// TIA Portal project "CHEMICAL DOSING PUMP" (V16)

(* hardware
DEVICE "S7-1200 station_1"  S7-1200 Station
   slot 0: "Rack_0"  S7-1200 Rack  Rack  V1.0
   slot 1: "PLC_1"  CPU 1214C DC/DC/DC  6ES7 214-1AG40-0XB0  V4.4
DEVICE "HMI_1"  TP900 Comfort
   slot 0: "HMI_1"  TP900 Comfort  6AV2 124-0JC01-0AX0  16.0.0.0
   slot 1: "HMI_RT_1"  TP900 Comfort  6AV2 124-0JC01-0AX0  16.0.0.0
   slot 5: "HMI_1.IE_CP_1"  PROFINET Interface  16.0.0.0
      slot 1: "PROFINET Interface_1"  PROFINET Interface
         slot 1: "Port_1"  Port
         slot 2: "Port_2"  Port
   slot 7: "HMI_1.MPI/DP_CP_1"  MPI/DP Interface  16.0.0.0
*)

// ===== PLC "PLC_1"  CPU 1214C DC/DC/DC =====

VAR_GLOBAL   // PLC tag table "Default tag table"
   "STOP SYSTEM" AT %M0.0 : Bool;
   "START SYSTEM" AT %M0.1 : Bool;
   "SYSTEM RUNNING" AT %M0.2 : Bool;
   "System_Byte" AT %MB2000 : Byte;
   "FirstScan" AT %M2000.0 : Bool;
   "DiagStatusUpdate" AT %M2000.1 : Bool;
   "AlwaysTRUE" AT %M2000.2 : Bool;
   "AlwaysFALSE" AT %M2000.3 : Bool;
   "System_Byte(1)" AT %MB1 : Byte;
   "Clock_Byte" AT %MB2001 : Byte;
   "Clock_10Hz" AT %M2001.0 : Bool;
   "Clock_5Hz" AT %M2001.1 : Bool;
   "Clock_2.5Hz" AT %M2001.2 : Bool;
   "Clock_2Hz" AT %M2001.3 : Bool;
   "Clock_1.25Hz" AT %M2001.4 : Bool;
   "Clock_1Hz" AT %M2001.5 : Bool;
   "Clock_0.625Hz" AT %M2001.6 : Bool;
   "Clock_0.5Hz" AT %M2001.7 : Bool;
   "TRIGGER 1" AT %M0.3 : Bool;
   "TRIGGER 2" AT %M0.4 : Bool;
   "DOSING PUMP 1" AT %Q0.0 : Bool;
   "HIGH LEVEL SET POINT" AT %MW4 : Int;
   "WATER TANK 2" AT %MW2 : Int;
   "TRIGGER 3" AT %M0.5 : Bool;
   "DOSING PUMP 2" AT %Q0.1 : Bool;
   "WATER TANK 2_2" AT %MW6 : Int;
   "TRIGGER 4" AT %M0.6 : Bool;
   "TRIGGER 5" AT %M0.7 : Bool;
   "TRIGGER 6" AT %M1.0 : Bool;
   "LOW LEVEL SETPOINT" AT %MW8 : Int;
END_VAR

// folder: System blocks/Program resources

DATA_BLOCK "C0"   // DB1
{ S7_Optimized_Access := 'TRUE' }
AUTHOR : Simatic
FAMILY : IEC
NAME : CNTR
VERSION : 1.0
// stored: InstanceOfName IEC_COUNTER
"IEC_COUNTER"
BEGIN
END_DATA_BLOCK

DATA_BLOCK "C1"   // DB2
{ S7_Optimized_Access := 'TRUE' }
AUTHOR : Simatic
FAMILY : IEC
NAME : CNTR
VERSION : 1.0
// stored: InstanceOfName IEC_COUNTER
"IEC_COUNTER"
BEGIN
END_DATA_BLOCK

// folder: (top level)

ORGANIZATION_BLOCK "Main"   // OB1, LAD, ProgramCycle
TITLE = "Main Program Sweep (Cycle)"
{ S7_Optimized_Access := 'TRUE' }
VERSION : 0.1
   VAR_INPUT
      Initial_Call : Bool;   // Initial call of this OB
      Remanence : Bool;   // =True, if remanent data are available
   END_VAR
   VAR_TEMP   // added for the SCL form of the ladder/FBD networks
      _w1 : Bool;
      _w2 : Bool;
      _w3 : Bool;
      _w4 : Bool;
   END_VAR
BEGIN

REGION Network 1: PROGRAM FOT STARTING AND STOPING A SYSTEM
   // * CREATING PROGRAM FOR STARTING AND STOPING CHEICAL DOSING SYSTEM
   // * ENABILY THE CLOCK MEMORY
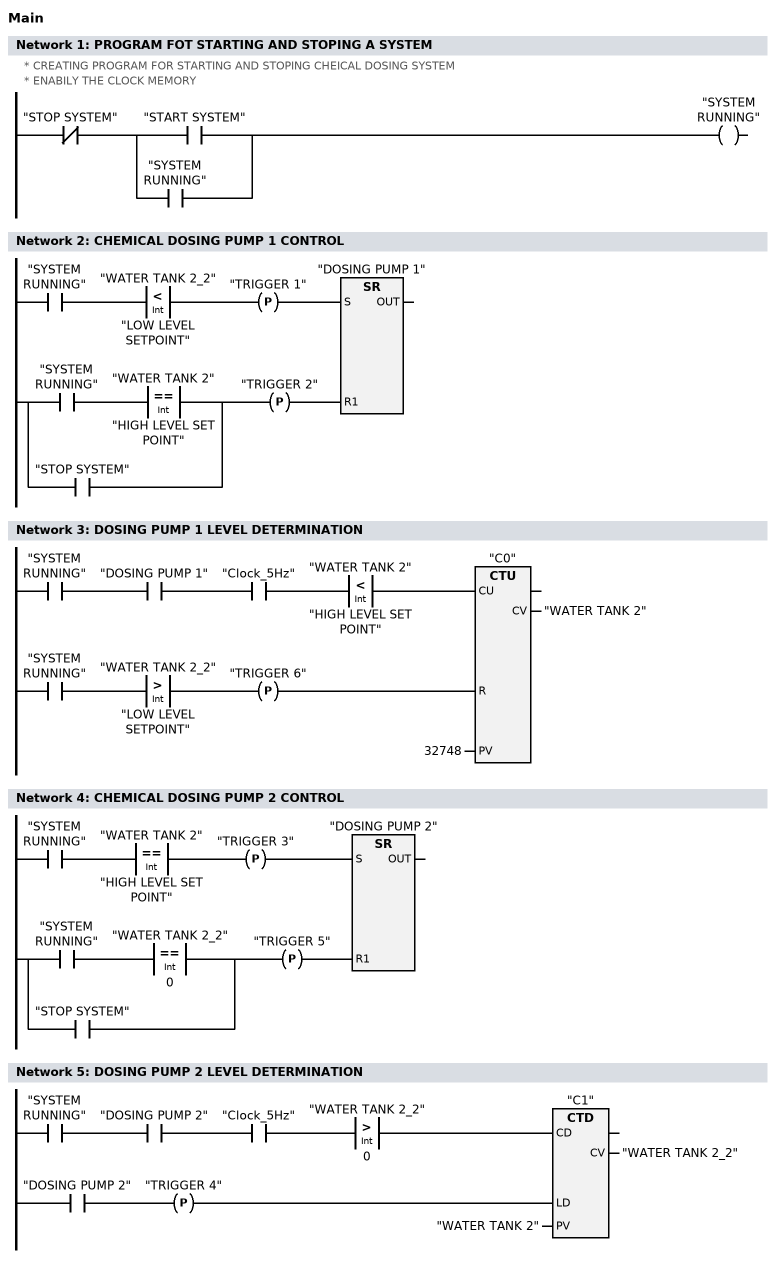
   RUNG wire#powerrail
      I_Contact( "STOP SYSTEM" )
      wire#w1
      Contact( "START SYSTEM" )
      wire#w2
      Coil( "SYSTEM RUNNING" )
   END_RUNG
   RUNG wire#w1
      Contact( "SYSTEM RUNNING" )
   END_RUNG wire#w2
   // the same network as SCL:
   "SYSTEM RUNNING" := NOT "STOP SYSTEM" AND ("START SYSTEM" OR "SYSTEM RUNNING");
END_REGION

REGION Network 2: CHEMICAL DOSING PUMP 1 CONTROL
   RUNG wire#powerrail
      Contact( "SYSTEM RUNNING" )
      { S7_Templates := "SrcType := Int" } LT_Contact(in1 := "WATER TANK 2_2", in2 := "LOW LEVEL SETPOINT")
      P_Trig( "TRIGGER 1" )
      S_SR(operand := "DOSING PUMP 1", r1 := wire#w2)
   END_RUNG
   RUNG wire#powerrail
      Contact( "SYSTEM RUNNING" )
      { S7_Templates := "SrcType := Int" } EQ_Contact(in1 := "WATER TANK 2", in2 := "HIGH LEVEL SET POINT")
      wire#w1
      P_Trig( "TRIGGER 2" )
   END_RUNG wire#w2
   RUNG wire#powerrail
      Contact( "STOP SYSTEM" )
   END_RUNG wire#w1
   // the same network as SCL:
   #_w1 := "SYSTEM RUNNING" AND ("WATER TANK 2_2" < "LOW LEVEL SETPOINT");
   #_w2 := #_w1 AND NOT "TRIGGER 1";   // rising edge
   "TRIGGER 1" := #_w1;
   #_w3 := ("SYSTEM RUNNING" AND ("WATER TANK 2" = "HIGH LEVEL SET POINT")) OR "STOP SYSTEM";
   #_w4 := #_w3 AND NOT "TRIGGER 2";   // rising edge
   "TRIGGER 2" := #_w3;
   IF #_w2 THEN
       "DOSING PUMP 1" := TRUE;   // SR flip-flop
   END_IF;
   IF #_w4 THEN "DOSING PUMP 1" := FALSE; END_IF;
END_REGION

REGION Network 3: DOSING PUMP 1 LEVEL DETERMINATION
   #_w1 := "SYSTEM RUNNING" AND ("WATER TANK 2_2" > "LOW LEVEL SETPOINT");
   #_w2 := #_w1 AND NOT "TRIGGER 6";   // rising edge
   "TRIGGER 6" := #_w1;
   "C0".CTU(CU := "SYSTEM RUNNING" AND "DOSING PUMP 1" AND "Clock_5Hz" AND ("WATER TANK 2" < "HIGH LEVEL SET POINT"),
            R := #_w2,
            PV := 32748,
            CV => "WATER TANK 2");
END_REGION

REGION Network 4: CHEMICAL DOSING PUMP 2 CONTROL
   RUNG wire#powerrail
      Contact( "SYSTEM RUNNING" )
      { S7_Templates := "SrcType := Int" } EQ_Contact(in1 := "WATER TANK 2", in2 := "HIGH LEVEL SET POINT")
      P_Trig( "TRIGGER 3" )
      S_SR(operand := "DOSING PUMP 2", r1 := wire#w2)
   END_RUNG
   RUNG wire#powerrail
      Contact( "SYSTEM RUNNING" )
      { S7_Templates := "SrcType := Int" } EQ_Contact(in1 := "WATER TANK 2_2", in2 := 0)
      wire#w1
      P_Trig( "TRIGGER 5" )
   END_RUNG wire#w2
   RUNG wire#powerrail
      Contact( "STOP SYSTEM" )
   END_RUNG wire#w1
   // the same network as SCL:
   #_w1 := "SYSTEM RUNNING" AND ("WATER TANK 2" = "HIGH LEVEL SET POINT");
   #_w2 := #_w1 AND NOT "TRIGGER 3";   // rising edge
   "TRIGGER 3" := #_w1;
   #_w3 := ("SYSTEM RUNNING" AND ("WATER TANK 2_2" = 0)) OR "STOP SYSTEM";
   #_w4 := #_w3 AND NOT "TRIGGER 5";   // rising edge
   "TRIGGER 5" := #_w3;
   IF #_w2 THEN
       "DOSING PUMP 2" := TRUE;   // SR flip-flop
   END_IF;
   IF #_w4 THEN "DOSING PUMP 2" := FALSE; END_IF;
END_REGION

REGION Network 5: DOSING PUMP 2 LEVEL DETERMINATION
   #_w1 := "DOSING PUMP 2" AND NOT "TRIGGER 4";   // rising edge
   "TRIGGER 4" := "DOSING PUMP 2";
   "C1".CTD(CD := "SYSTEM RUNNING" AND "DOSING PUMP 2" AND "Clock_5Hz" AND ("WATER TANK 2_2" > 0),
            LD := #_w1,
            PV := "WATER TANK 2",
            CV => "WATER TANK 2_2");
END_REGION
END_ORGANIZATION_BLOCK

(* ===== HMI "HMI_RT_1" =====
system functions are stored by id; their names below are inferred from use
connection "HMI_Connection_1": ETHERNET, S7_1200_OMS

HMI tags "Default tag table"
   "Tag_ScreenNumber" : UInt, internal
   "WATER TANK 2" : Int = PLC "WATER TANK 2" AT %MW2, 1 s
   "WATER TANK 2_2" : Int = PLC "WATER TANK 2_2" AT %MW6, 1 s
   "START SYSTEM" : Bool = PLC "STOP SYSTEM" AT %M0.0, 1 s
   "STOP SYSTEM" : Bool = PLC "START SYSTEM" AT %M0.1, 1 s
   "DOSING PUMP 1" : Bool = PLC "DOSING PUMP 1" AT %Q0.0, 1 s
   "DOSING PUMP 2" : Bool = PLC "DOSING PUMP 2" AT %Q0.1, 1 s
   "LOW LEVEL SETPOINT" : Int = PLC "LOW LEVEL SETPOINT" AT %MW8, 1 s
   "HIGH LEVEL SET POINT" : Int = PLC "HIGH LEVEL SET POINT" AT %MW4, 1 s
   "SYSTEM RUNNING" : Bool = PLC "SYSTEM RUNNING" AT %M0.2, 1 s

screen "Root screen" 800x420, template "Template_1"
   on GenerateScreen: SetTag("Tag_ScreenNumber", 1)
   SymbolLibrary "Symbol library_1" at 626,75 size 164x120
      Appearance <- "DOSING PUMP 1"
   SymbolLibrary "Symbol library_2" at 36,242 size 187x102
      Appearance <- "DOSING PUMP 2"
   SymbolLibrary "Symbol library_3" at 503,134 size 127x35
      Appearance <- "DOSING PUMP 1"
   SymbolLibrary "Symbol library_4" at 446,134 size 60x68
      Appearance <- "DOSING PUMP 1"
   SymbolLibrary "Symbol library_5" at 446,200 size 31x82
      Appearance <- "DOSING PUMP 1"
   SymbolLibrary "Symbol library_9" at 627,11 size 41x67
      Appearance <- "DOSING PUMP 1"
   SymbolLibrary "Symbol library_10" at 222,278 size 52x46
      Appearance <- "DOSING PUMP 2"
   SymbolLibrary "Symbol library_11" at 248,193 size 26x94
      Appearance <- "DOSING PUMP 2"
   SymbolLibrary "Symbol library_12" at 159,209 size 39x37
      Appearance <- "DOSING PUMP 2"
   SymbolLibrary "Symbol library_13" at 27,208 size 138x21
      Appearance <- "DOSING PUMP 2"
   Bar "Bar_2" at 52,76 size 280x126; MinimumValue 0; MaximumValue 250
      ProcessValue <- "WATER TANK 2_2"
      Visibility <- "DOSING PUMP 1"
   TextField "Text field_1" at 607,218 size 161x25; Text 'CONTROL PANEL'
   Circle "Circle_1" at 648,251 size 48x48
      Appearance <- "SYSTEM RUNNING"
   TextField "Text field_2" at 667,85 size 145x22; Text 'FILLING PUMP 1'
   TextField "Text field_3" at 13,255 size 154x22; Text 'DOSSING PUMP 2'
   SymbolLibrary "Symbol library_6" at 164,11 size 465x32
      Appearance <- "DOSING PUMP 1"
   IOField "I/O field_1" at 335,176 size 52x29; FormatPattern 999
      ProcessValue <- "LOW LEVEL SETPOINT"
   IOField "I/O field_2" at 334,85 size 52x29; FormatPattern 999
      ProcessValue <- "HIGH LEVEL SET POINT"
   TextField "Text field_4" at 384,90 size 21x25; Text 'M'
   TextField "Text field_5" at 386,179 size 21x25; Text 'M'
   Bar "Bar_1" at 53,77 size 280x125; MinimumValue 0; MaximumValue 250
      ProcessValue <- "WATER TANK 2"
      Visibility <- "DOSING PUMP 2"
   SymbolLibrary "Symbol library_7" at 115,10 size 50x66
      Appearance <- "DOSING PUMP 1"
   SymbolLibrary "Symbol library_8" at 115,68 size 26x43
      Appearance <- "DOSING PUMP 1"
   Button "Button_1" at 588,304 size 68x28; TextOff 'START'
      on Press: function_b14e0dd5("STOP SYSTEM", 0)
   Button "Button_2" at 718,306 size 68x28; TextOff 'STOP'
      on Press: function_b14e0dd5("START SYSTEM", 0)
   TextField "Text field_6" at 360,304 size 228x25; Text 'CHEMICAL RESERVOUR'
   TextField "Text field_7" at 148,168 size 134x25; Text 'FEED HOPPER'

Template "Template_1" 800x420
   Button "Exit" at 720,360 size 78x58; TextOff 'Exit'; PictureOff "ExitRuntime_TP900_Comfort_TR"; PictureOn "ExitRuntime_TP900_Comfort_TR"
      on Release: StopRuntime(0)
   Button "Template_Button" at 640,360 size 78x58; TextOff 'Text'
   Button "Template_Button_1" at 560,360 size 78x58; TextOff 'Text'
   Button "Template_Button_2" at 480,360 size 78x58; TextOff 'Text'
   Button "Template_Button_3" at 400,360 size 78x58; TextOff 'Text'
   Button "Template_Button_4" at 321,360 size 78x58; TextOff 'Text'
   Button "Template_Button_5" at 241,360 size 78x58; TextOff 'Text'
   Button "Template_Button_6" at 161,360 size 78x58; TextOff 'Text'
   Button "Alarms" at 81,360 size 78x58; TextOff 'Alarms'; PictureOff "AlarmDisplay_TP900_Comfort_TR"; PictureOn "AlarmDisplay_TP900_Comfort_TR"
      on Release: function_ef3f5d25("Alarm window_Unacknowledged", -1)
   Button "Start screen" at 1,360 size 78x58; TextOff 'Start screen'; PictureOff "NavigateHome_TP900_Comfort_TR"; PictureOn "NavigateHome_TP900_Comfort_TR"
      on Release: ActivateScreen("Root screen", 0)
*)